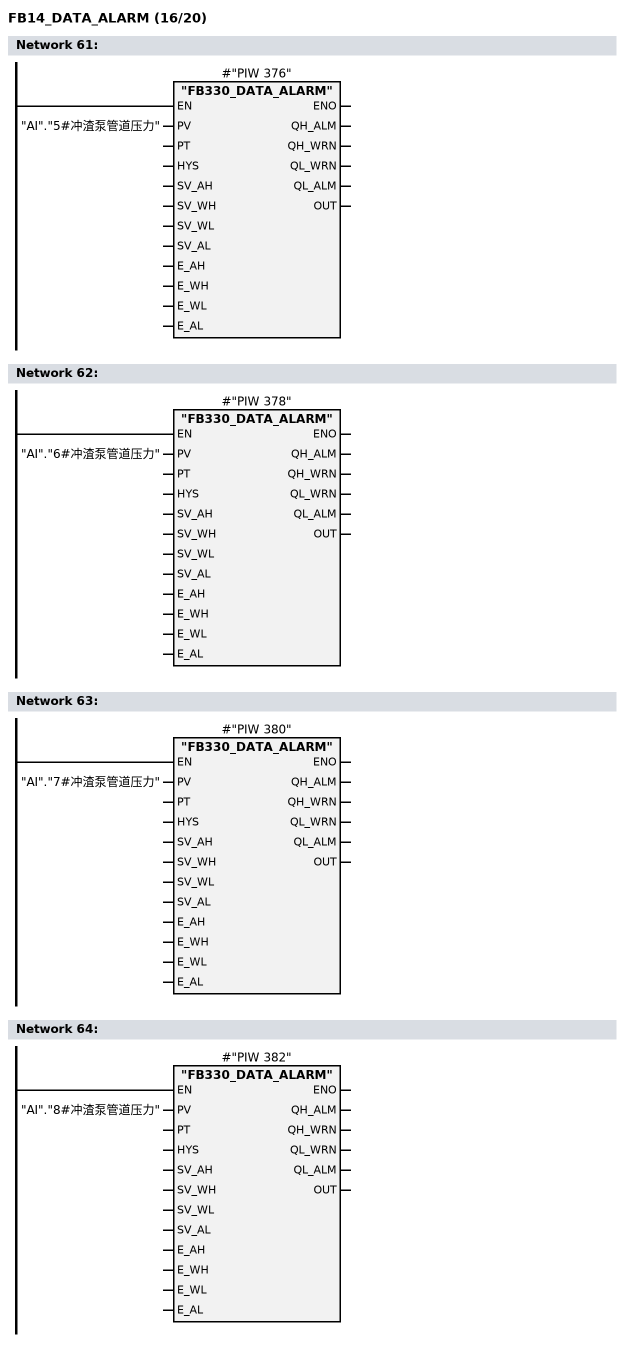
   RUNG wire#powerrail
      #"PIW 376"(PV := "AI"."5#冲渣泵管道压力", PT :=, HYS :=, SV_AH :=, SV_WH :=, SV_WL :=, SV_AL :=, E_AH :=, E_WH :=, E_WL :=, E_AL :=, QH_ALM =>, QH_WRN =>, QL_WRN =>, QL_ALM =>, OUT =>)
   END_RUNG
   // the same network as SCL:
   #"PIW 376"(PV := "AI"."5#冲渣泵管道压力");   // "FB330_DATA_ALARM"
END_REGION

REGION Network 62
   RUNG wire#powerrail
      #"PIW 378"(PV := "AI"."6#冲渣泵管道压力", PT :=, HYS :=, SV_AH :=, SV_WH :=, SV_WL :=, SV_AL :=, E_AH :=, E_WH :=, E_WL :=, E_AL :=, QH_ALM =>, QH_WRN =>, QL_WRN =>, QL_ALM =>, OUT =>)
   END_RUNG
   // the same network as SCL:
   #"PIW 378"(PV := "AI"."6#冲渣泵管道压力");   // "FB330_DATA_ALARM"
END_REGION

REGION Network 63
   RUNG wire#powerrail
      #"PIW 380"(PV := "AI"."7#冲渣泵管道压力", PT :=, HYS :=, SV_AH :=, SV_WH :=, SV_WL :=, SV_AL :=, E_AH :=, E_WH :=, E_WL :=, E_AL :=, QH_ALM =>, QH_WRN =>, QL_WRN =>, QL_ALM =>, OUT =>)
   END_RUNG
   // the same network as SCL:
   #"PIW 380"(PV := "AI"."7#冲渣泵管道压力");   // "FB330_DATA_ALARM"
END_REGION

REGION Network 64
   RUNG wire#powerrail
      #"PIW 382"(PV := "AI"."8#冲渣泵管道压力", PT :=, HYS :=, SV_AH :=, SV_WH :=, SV_WL :=, SV_AL :=, E_AH :=, E_WH :=, E_WL :=, E_AL :=, QH_ALM =>, QH_WRN =>, QL_WRN =>, QL_ALM =>, OUT =>)
   END_RUNG
   // the same network as SCL:
   #"PIW 382"(PV := "AI"."8#冲渣泵管道压力");   // "FB330_DATA_ALARM"
END_REGION

REGION Network 65
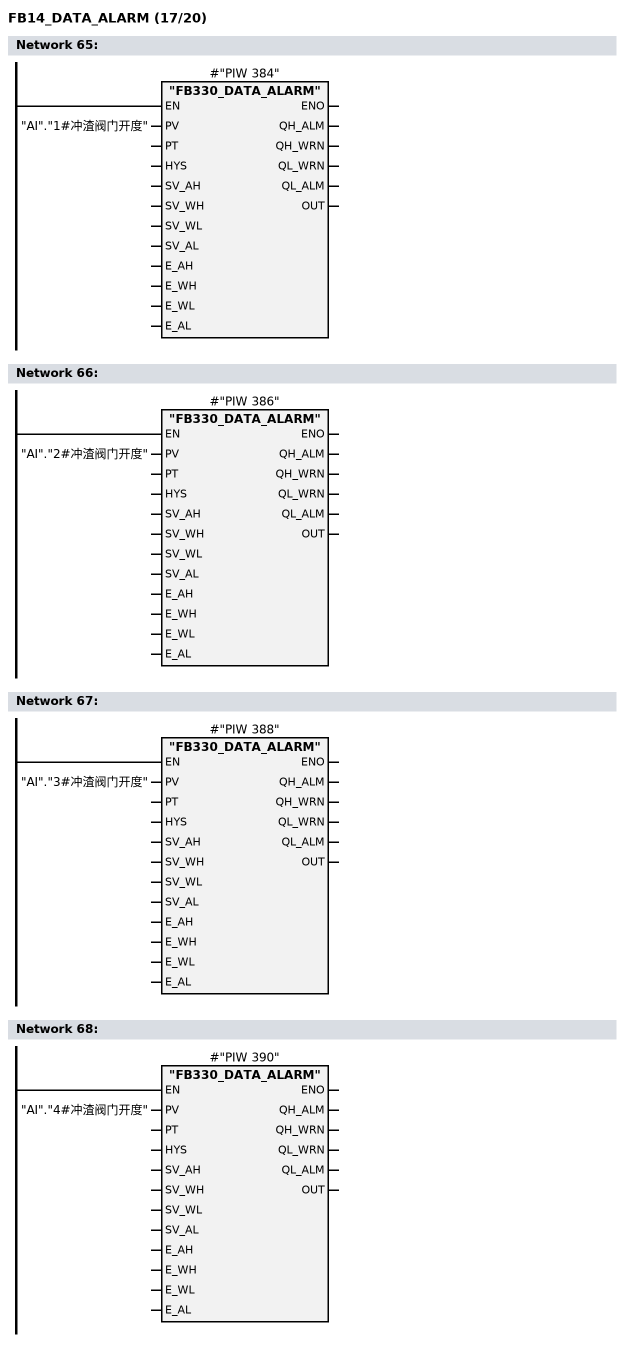
   RUNG wire#powerrail
      #"PIW 384"(PV := "AI"."1#冲渣阀门开度", PT :=, HYS :=, SV_AH :=, SV_WH :=, SV_WL :=, SV_AL :=, E_AH :=, E_WH :=, E_WL :=, E_AL :=, QH_ALM =>, QH_WRN =>, QL_WRN =>, QL_ALM =>, OUT =>)
   END_RUNG
   // the same network as SCL:
   #"PIW 384"(PV := "AI"."1#冲渣阀门开度");   // "FB330_DATA_ALARM"
END_REGION

REGION Network 66
   RUNG wire#powerrail
      #"PIW 386"(PV := "AI"."2#冲渣阀门开度", PT :=, HYS :=, SV_AH :=, SV_WH :=, SV_WL :=, SV_AL :=, E_AH :=, E_WH :=, E_WL :=, E_AL :=, QH_ALM =>, QH_WRN =>, QL_WRN =>, QL_ALM =>, OUT =>)
   END_RUNG
   // the same network as SCL:
   #"PIW 386"(PV := "AI"."2#冲渣阀门开度");   // "FB330_DATA_ALARM"
END_REGION

REGION Network 67
   RUNG wire#powerrail
      #"PIW 388"(PV := "AI"."3#冲渣阀门开度", PT :=, HYS :=, SV_AH :=, SV_WH :=, SV_WL :=, SV_AL :=, E_AH :=, E_WH :=, E_WL :=, E_AL :=, QH_ALM =>, QH_WRN =>, QL_WRN =>, QL_ALM =>, OUT =>)
   END_RUNG
   // the same network as SCL:
   #"PIW 388"(PV := "AI"."3#冲渣阀门开度");   // "FB330_DATA_ALARM"
END_REGION

REGION Network 68
   RUNG wire#powerrail
      #"PIW 390"(PV := "AI"."4#冲渣阀门开度", PT :=, HYS :=, SV_AH :=, SV_WH :=, SV_WL :=, SV_AL :=, E_AH :=, E_WH :=, E_WL :=, E_AL :=, QH_ALM =>, QH_WRN =>, QL_WRN =>, QL_ALM =>, OUT =>)
   END_RUNG
   // the same network as SCL:
   #"PIW 390"(PV := "AI"."4#冲渣阀门开度");   // "FB330_DATA_ALARM"
END_REGION

REGION Network 69
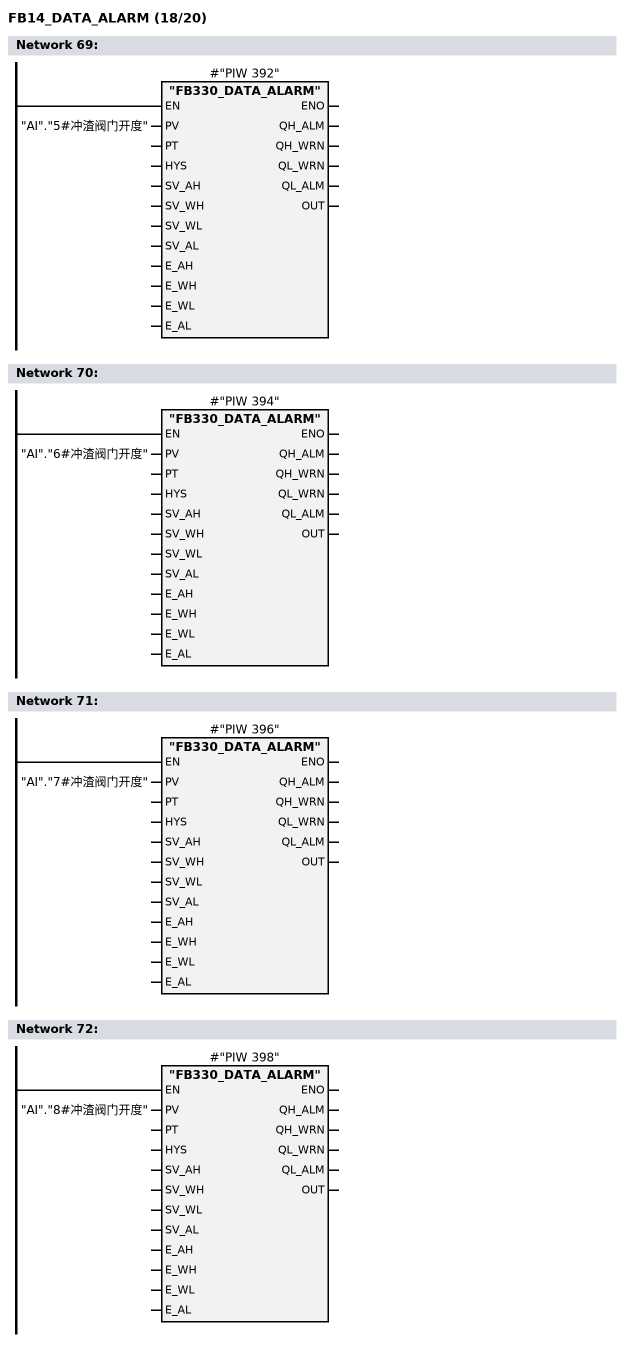
   RUNG wire#powerrail
      #"PIW 392"(PV := "AI"."5#冲渣阀门开度", PT :=, HYS :=, SV_AH :=, SV_WH :=, SV_WL :=, SV_AL :=, E_AH :=, E_WH :=, E_WL :=, E_AL :=, QH_ALM =>, QH_WRN =>, QL_WRN =>, QL_ALM =>, OUT =>)
   END_RUNG
   // the same network as SCL:
   #"PIW 392"(PV := "AI"."5#冲渣阀门开度");   // "FB330_DATA_ALARM"
END_REGION

REGION Network 70
   RUNG wire#powerrail
      #"PIW 394"(PV := "AI"."6#冲渣阀门开度", PT :=, HYS :=, SV_AH :=, SV_WH :=, SV_WL :=, SV_AL :=, E_AH :=, E_WH :=, E_WL :=, E_AL :=, QH_ALM =>, QH_WRN =>, QL_WRN =>, QL_ALM =>, OUT =>)
   END_RUNG
   // the same network as SCL:
   #"PIW 394"(PV := "AI"."6#冲渣阀门开度");   // "FB330_DATA_ALARM"
END_REGION

REGION Network 71
   RUNG wire#powerrail
      #"PIW 396"(PV := "AI"."7#冲渣阀门开度", PT :=, HYS :=, SV_AH :=, SV_WH :=, SV_WL :=, SV_AL :=, E_AH :=, E_WH :=, E_WL :=, E_AL :=, QH_ALM =>, QH_WRN =>, QL_WRN =>, QL_ALM =>, OUT =>)
   END_RUNG
   // the same network as SCL:
   #"PIW 396"(PV := "AI"."7#冲渣阀门开度");   // "FB330_DATA_ALARM"
END_REGION

REGION Network 72
   RUNG wire#powerrail
      #"PIW 398"(PV := "AI"."8#冲渣阀门开度", PT :=, HYS :=, SV_AH :=, SV_WH :=, SV_WL :=, SV_AL :=, E_AH :=, E_WH :=, E_WL :=, E_AL :=, QH_ALM =>, QH_WRN =>, QL_WRN =>, QL_ALM =>, OUT =>)
   END_RUNG
   // the same network as SCL:
   #"PIW 398"(PV := "AI"."8#冲渣阀门开度");   // "FB330_DATA_ALARM"
END_REGION

REGION Network 73
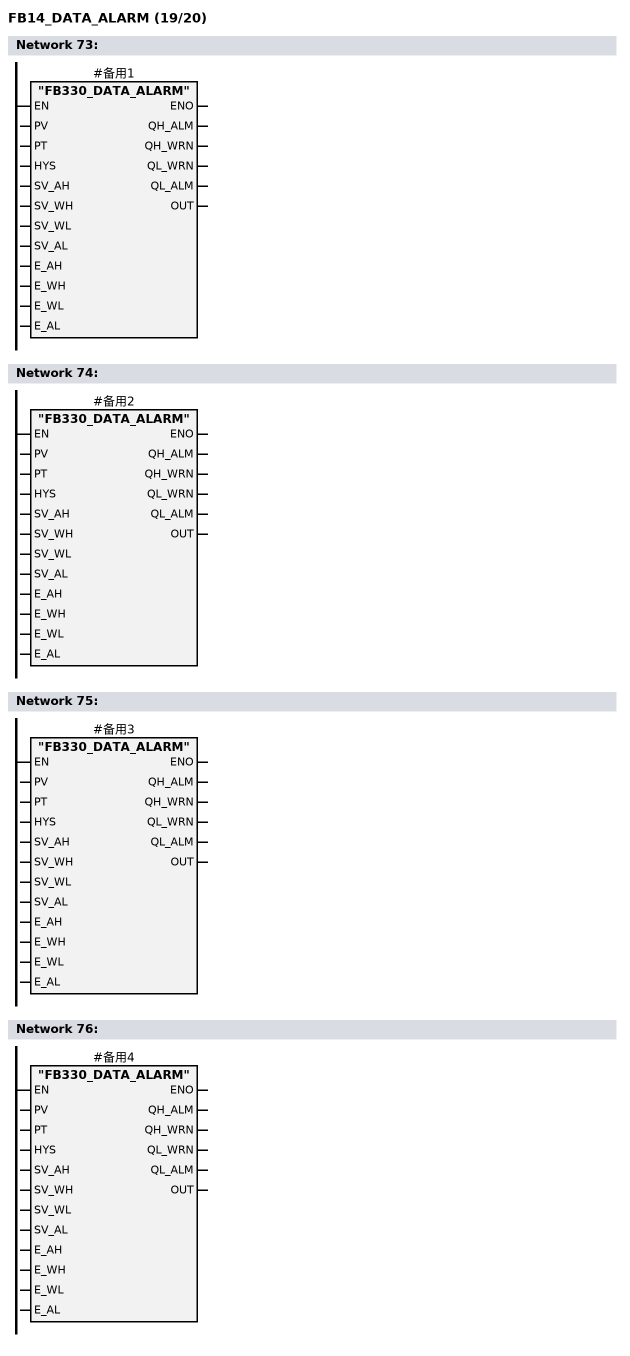
   RUNG wire#powerrail
      #备用1(PV :=, PT :=, HYS :=, SV_AH :=, SV_WH :=, SV_WL :=, SV_AL :=, E_AH :=, E_WH :=, E_WL :=, E_AL :=, QH_ALM =>, QH_WRN =>, QL_WRN =>, QL_ALM =>, OUT =>)
   END_RUNG
   // the same network as SCL:
   #备用1();   // "FB330_DATA_ALARM"
END_REGION

REGION Network 74
   RUNG wire#powerrail
      #备用2(PV :=, PT :=, HYS :=, SV_AH :=, SV_WH :=, SV_WL :=, SV_AL :=, E_AH :=, E_WH :=, E_WL :=, E_AL :=, QH_ALM =>, QH_WRN =>, QL_WRN =>, QL_ALM =>, OUT =>)
   END_RUNG
   // the same network as SCL:
   #备用2();   // "FB330_DATA_ALARM"
END_REGION

REGION Network 75
   RUNG wire#powerrail
      #备用3(PV :=, PT :=, HYS :=, SV_AH :=, SV_WH :=, SV_WL :=, SV_AL :=, E_AH :=, E_WH :=, E_WL :=, E_AL :=, QH_ALM =>, QH_WRN =>, QL_WRN =>, QL_ALM =>, OUT =>)
   END_RUNG
   // the same network as SCL:
   #备用3();   // "FB330_DATA_ALARM"
END_REGION

REGION Network 76
   RUNG wire#powerrail
      #备用4(PV :=, PT :=, HYS :=, SV_AH :=, SV_WH :=, SV_WL :=, SV_AL :=, E_AH :=, E_WH :=, E_WL :=, E_AL :=, QH_ALM =>, QH_WRN =>, QL_WRN =>, QL_ALM =>, OUT =>)
   END_RUNG
   // the same network as SCL:
   #备用4();   // "FB330_DATA_ALARM"
END_REGION

REGION Network 77
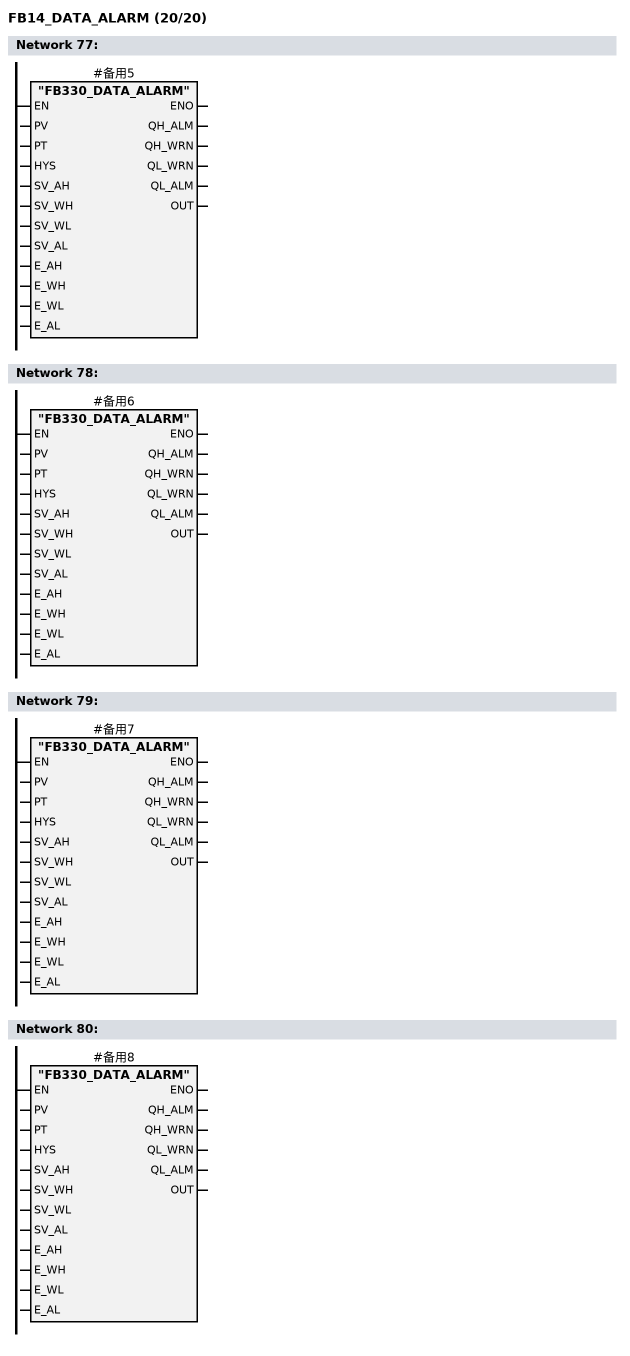
   RUNG wire#powerrail
      #备用5(PV :=, PT :=, HYS :=, SV_AH :=, SV_WH :=, SV_WL :=, SV_AL :=, E_AH :=, E_WH :=, E_WL :=, E_AL :=, QH_ALM =>, QH_WRN =>, QL_WRN =>, QL_ALM =>, OUT =>)
   END_RUNG
   // the same network as SCL:
   #备用5();   // "FB330_DATA_ALARM"
END_REGION

REGION Network 78
   RUNG wire#powerrail
      #备用6(PV :=, PT :=, HYS :=, SV_AH :=, SV_WH :=, SV_WL :=, SV_AL :=, E_AH :=, E_WH :=, E_WL :=, E_AL :=, QH_ALM =>, QH_WRN =>, QL_WRN =>, QL_ALM =>, OUT =>)
   END_RUNG
   // the same network as SCL:
   #备用6();   // "FB330_DATA_ALARM"
END_REGION

REGION Network 79
   RUNG wire#powerrail
      #备用7(PV :=, PT :=, HYS :=, SV_AH :=, SV_WH :=, SV_WL :=, SV_AL :=, E_AH :=, E_WH :=, E_WL :=, E_AL :=, QH_ALM =>, QH_WRN =>, QL_WRN =>, QL_ALM =>, OUT =>)
   END_RUNG
   // the same network as SCL:
   #备用7();   // "FB330_DATA_ALARM"
END_REGION

REGION Network 80
   RUNG wire#powerrail
      #备用8(PV :=, PT :=, HYS :=, SV_AH :=, SV_WH :=, SV_WL :=, SV_AL :=, E_AH :=, E_WH :=, E_WL :=, E_AL :=, QH_ALM =>, QH_WRN =>, QL_WRN =>, QL_ALM =>, OUT =>)
   END_RUNG
   // the same network as SCL:
   #备用8();   // "FB330_DATA_ALARM"
END_REGION
END_FUNCTION_BLOCK

FUNCTION_BLOCK "FB15_MOTOR_AUTO-st"   // FB15, LAD
{ S7_Optimized_Access := 'FALSE' }
VERSION : 0.1
   VAR
      "1#冲渣泵驱动" : "FB310_MOTOR_AUTO_ST_model";
      "2#冲渣泵驱动" : "FB310_MOTOR_AUTO_ST_model";
      "3#冲渣泵驱动" : "FB310_MOTOR_AUTO_ST_model";
      "4#冲渣泵驱动" : "FB310_MOTOR_AUTO_ST_model";
      "5#冲渣泵驱动" : "FB310_MOTOR_AUTO_ST_model";
      "6#冲渣泵驱动" : "FB310_MOTOR_AUTO_ST_model";
      "7#冲渣泵驱动" : "FB310_MOTOR_AUTO_ST_model";
      "8#冲渣泵驱动" : "FB310_MOTOR_AUTO_ST_model";
      "1#浊环热水泵驱动" : "FB310_MOTOR_AUTO_ST_model";
      "2#浊环热水泵驱动" : "FB310_MOTOR_AUTO_ST_model";
      "3#浊环热水泵驱动" : "FB310_MOTOR_AUTO_ST_model";
      "4#浊环热水泵驱动" : "FB310_MOTOR_AUTO_ST_model";
      "5#浊环热水泵驱动" : "FB310_MOTOR_AUTO_ST_model";
      "6#浊环热水泵驱动" : "FB310_MOTOR_AUTO_ST_model";
      "7#浊环热水泵驱动" : "FB310_MOTOR_AUTO_ST_model";
      "8#浊环热水泵驱动" : "FB310_MOTOR_AUTO_ST_model";
      "1#炉体循环水泵驱动" : "FB310_MOTOR_AUTO_ST_model";
      "2#炉体循环水泵驱动" : "FB310_MOTOR_AUTO_ST_model";
      "3#炉体循环水泵驱动" : "FB310_MOTOR_AUTO_ST_model";
      "1#电极循环水泵驱动" : "FB310_MOTOR_AUTO_ST_model";
      "2#电极循环水泵驱动" : "FB310_MOTOR_AUTO_ST_model";
      "3#电极循环水泵驱动" : "FB310_MOTOR_AUTO_ST_model";
      "4#电极循环水泵驱动" : "FB310_MOTOR_AUTO_ST_model";
      "1#净环热水泵驱动" : "FB310_MOTOR_AUTO_ST_model";
      "2#净环热水泵驱动" : "FB310_MOTOR_AUTO_ST_model";
      "3#净环热水泵驱动" : "FB310_MOTOR_AUTO_ST_model";
      "4#净环热水泵驱动" : "FB310_MOTOR_AUTO_ST_model";
      "5#净环热水泵驱动" : "FB310_MOTOR_AUTO_ST_model";
      "1#柴油泵驱动" : "FB310_MOTOR_AUTO_ST_model";
      "2#柴油泵驱动" : "FB310_MOTOR_AUTO_ST_model";
      窑冷却泵驱动 : "FB310_MOTOR_AUTO_ST_model";
      Static1 : "FB310_MOTOR_AUTO_ST_model";
      Static2 : "FB310_MOTOR_AUTO_ST_model";
      Static3 : "FB310_MOTOR_AUTO_ST_model";
      Static4 : "FB310_MOTOR_AUTO_ST_model";
      Static5 : "FB310_MOTOR_AUTO_ST_model";
      Static6 : "FB310_MOTOR_AUTO_ST_model";
      Static7 : "FB310_MOTOR_AUTO_ST_model";
      Static8 : "FB310_MOTOR_AUTO_ST_model";
      Static9 : "FB310_MOTOR_AUTO_ST_model";
      Static10 : "FB310_MOTOR_AUTO_ST_model";
   END_VAR
BEGIN

REGION Network 1
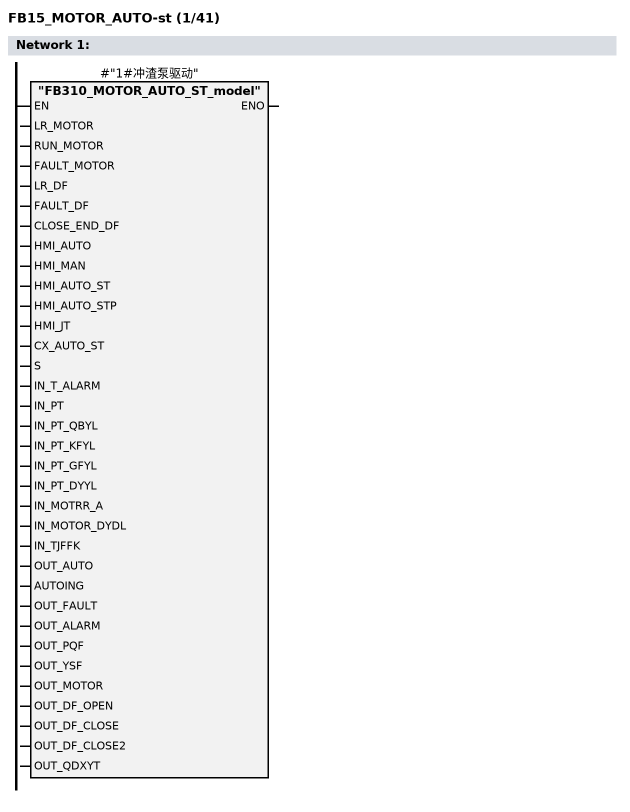
   RUNG wire#powerrail
      #"1#冲渣泵驱动"(LR_MOTOR :=, RUN_MOTOR :=, FAULT_MOTOR :=, LR_DF :=, FAULT_DF :=, CLOSE_END_DF :=, HMI_AUTO :=, HMI_MAN :=, HMI_AUTO_ST :=, HMI_AUTO_STP :=, HMI_JT :=, CX_AUTO_ST :=, S :=, IN_T_ALARM :=, IN_PT :=, IN_PT_QBYL :=, IN_PT_KFYL :=, IN_PT_GFYL :=, IN_PT_DYYL :=, IN_MOTRR_A :=, IN_MOTOR_DYDL :=, IN_TJFFK :=, OUT_AUTO :=, AUTOING :=, OUT_FAULT :=, OUT_ALARM :=, OUT_PQF :=, OUT_YSF :=, OUT_MOTOR :=, OUT_DF_OPEN :=, OUT_DF_CLOSE :=, OUT_DF_CLOSE2 :=, OUT_QDXYT :=)
   END_RUNG
   // the same network as SCL:
   #"1#冲渣泵驱动"();   // "FB310_MOTOR_AUTO_ST_model"
END_REGION

REGION Network 2
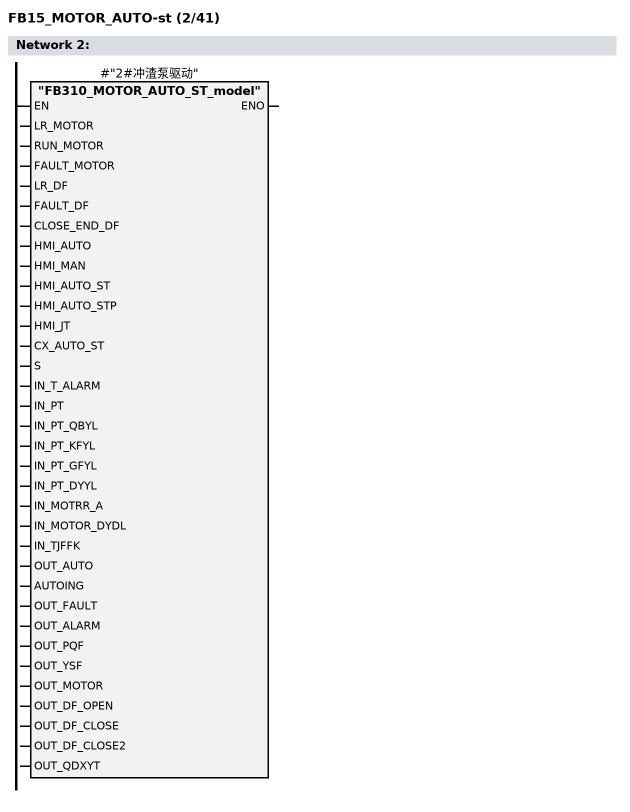
   RUNG wire#powerrail
      #"2#冲渣泵驱动"(LR_MOTOR :=, RUN_MOTOR :=, FAULT_MOTOR :=, LR_DF :=, FAULT_DF :=, CLOSE_END_DF :=, HMI_AUTO :=, HMI_MAN :=, HMI_AUTO_ST :=, HMI_AUTO_STP :=, HMI_JT :=, CX_AUTO_ST :=, S :=, IN_T_ALARM :=, IN_PT :=, IN_PT_QBYL :=, IN_PT_KFYL :=, IN_PT_GFYL :=, IN_PT_DYYL :=, IN_MOTRR_A :=, IN_MOTOR_DYDL :=, IN_TJFFK :=, OUT_AUTO :=, AUTOING :=, OUT_FAULT :=, OUT_ALARM :=, OUT_PQF :=, OUT_YSF :=, OUT_MOTOR :=, OUT_DF_OPEN :=, OUT_DF_CLOSE :=, OUT_DF_CLOSE2 :=, OUT_QDXYT :=)
   END_RUNG
   // the same network as SCL:
   #"2#冲渣泵驱动"();   // "FB310_MOTOR_AUTO_ST_model"
END_REGION

REGION Network 3
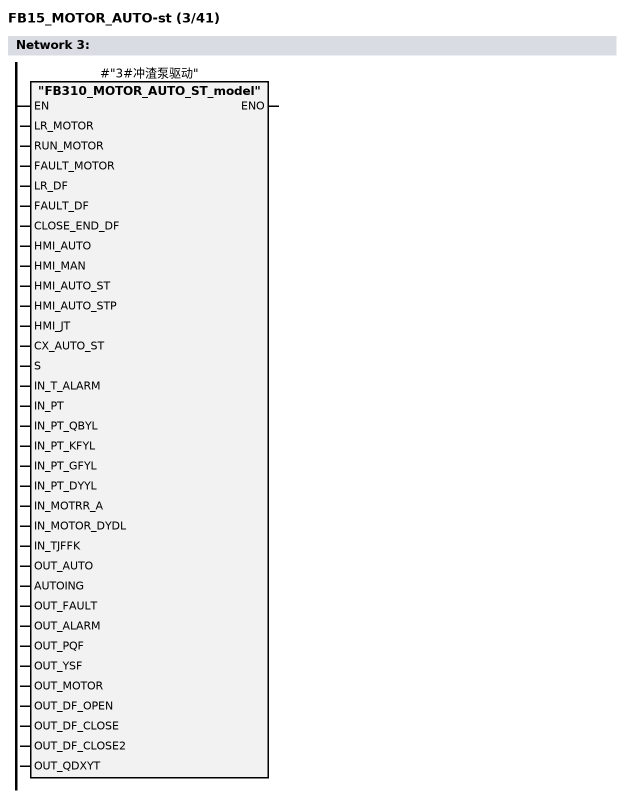
   RUNG wire#powerrail
      #"3#冲渣泵驱动"(LR_MOTOR :=, RUN_MOTOR :=, FAULT_MOTOR :=, LR_DF :=, FAULT_DF :=, CLOSE_END_DF :=, HMI_AUTO :=, HMI_MAN :=, HMI_AUTO_ST :=, HMI_AUTO_STP :=, HMI_JT :=, CX_AUTO_ST :=, S :=, IN_T_ALARM :=, IN_PT :=, IN_PT_QBYL :=, IN_PT_KFYL :=, IN_PT_GFYL :=, IN_PT_DYYL :=, IN_MOTRR_A :=, IN_MOTOR_DYDL :=, IN_TJFFK :=, OUT_AUTO :=, AUTOING :=, OUT_FAULT :=, OUT_ALARM :=, OUT_PQF :=, OUT_YSF :=, OUT_MOTOR :=, OUT_DF_OPEN :=, OUT_DF_CLOSE :=, OUT_DF_CLOSE2 :=, OUT_QDXYT :=)
   END_RUNG
   // the same network as SCL:
   #"3#冲渣泵驱动"();   // "FB310_MOTOR_AUTO_ST_model"
END_REGION

REGION Network 4
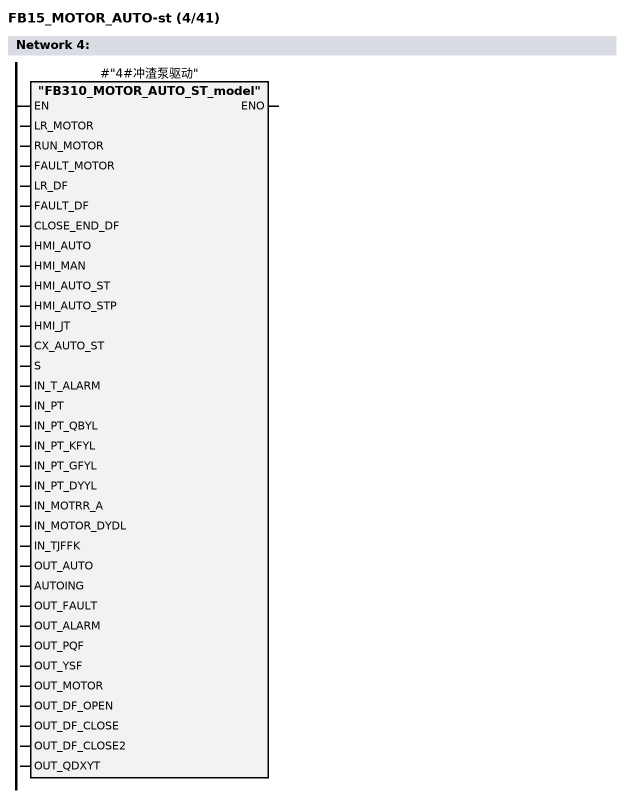
   RUNG wire#powerrail
      #"4#冲渣泵驱动"(LR_MOTOR :=, RUN_MOTOR :=, FAULT_MOTOR :=, LR_DF :=, FAULT_DF :=, CLOSE_END_DF :=, HMI_AUTO :=, HMI_MAN :=, HMI_AUTO_ST :=, HMI_AUTO_STP :=, HMI_JT :=, CX_AUTO_ST :=, S :=, IN_T_ALARM :=, IN_PT :=, IN_PT_QBYL :=, IN_PT_KFYL :=, IN_PT_GFYL :=, IN_PT_DYYL :=, IN_MOTRR_A :=, IN_MOTOR_DYDL :=, IN_TJFFK :=, OUT_AUTO :=, AUTOING :=, OUT_FAULT :=, OUT_ALARM :=, OUT_PQF :=, OUT_YSF :=, OUT_MOTOR :=, OUT_DF_OPEN :=, OUT_DF_CLOSE :=, OUT_DF_CLOSE2 :=, OUT_QDXYT :=)
   END_RUNG
   // the same network as SCL:
   #"4#冲渣泵驱动"();   // "FB310_MOTOR_AUTO_ST_model"
END_REGION

REGION Network 5